   "102_Pilot_Burner_DB_FD_VRFCTN_TMR_ET" : Time = PLC "102_Pilot_Burner_DB".FD_VRFCTN_TMR.ET, 1 s
   "102_Pilot_Burner_DB_FD_VRFCTN_TMR II_ET" : Time = PLC "20_TANKS_IP_DATA".RIO_02.SECOND_TANK.BWT_DO, 1 s
   "86_Times_PIT358 Delay" : Time = PLC "86_Times"."PIT358 Delay", 1 s
   "86_Times_PIT348 Delay" : Time = PLC "86_Times"."PIT348 Delay", 1 s
   "PGC Flush_DB_Temperature Setpoint" : Real = PLC "PGC Flush_DB"."Temperature Setpoint", 1 s
   "2062_Warning_Data_Water Level Override" : Bool = PLC "2062_Warning_Data"."Water Level Override" AT %DB2062.DBX376.0, 1 s
   "2062_Warning_Data_Water Level Override_Aux" : Bool = PLC "2062_Warning_Data"."Water Level Override_Aux" AT %DB2062.DBX376.2, 1 s
   "Sequence Times_DB_Boost" : Bool = PLC "Sequence Times_DB".Boost, 1 s
   "86_Times_FS320 delay" : Time = PLC "86_Times"."FS320 delay", 1 s
   "86_Times_FS317 delay" : Time = PLC "86_Times"."FS317 delay", 1 s
   "86_Times_PS101 Alarm Delay" : Time = PLC "86_Times"."PS101 Alarm Delay", 1 s
   "82_To_HMI_FS350 Animation" : Int = PLC "82_To_HMI"."FS350 Animation", 1 s
   "82_To_HMI_FS332 Animation" : Int = PLC "82_To_HMI"."FS332 Animation", 1 s
   "82_To_HMI_P304 Animation" : Int = PLC "82_To_HMI"."P304 Animation", 1 s
   "Sequence Times_DB_Post-Dwell Timer_Q" : Bool = PLC "Sequence Times_DB"."Post-Dwell Timer".Q, 1 s
      on ChangeValue: "TreatmentCycleCompleted"()
   "51_SLAVE_STATUS_MAIN_BURNER_ACTV" : Bool = PLC "51_SLAVE_STATUS".MAIN_BURNER_ACTV AT %DB51.DBX17.5, 1 s
   "Main Burner Animation_DB_Animation" : Int = PLC "Main Burner Animation_DB".Animation, 1 s
   "20_TANKS_IP_DATA_RIO_01_FIRST_TANK_USD FLOW  N" : Real = PLC "20_TANKS_IP_DATA".RIO_01.FIRST_TANK."USD FLOW  N", 1 s
   "20_TANKS_IP_DATA_RIO_01_FIRST_TANK_MBG_FLOW N" : Real = PLC "20_TANKS_IP_DATA".RIO_01.FIRST_TANK."MBG_FLOW N", 1 s
   "20_TANKS_IP_DATA_RIO_01_SECOND_TANK_MBG_FLOW N" : Real = PLC "20_TANKS_IP_DATA".RIO_01.SECOND_TANK."MBG_FLOW N", 1 s
   "20_TANKS_IP_DATA_RIO_01_SECOND_TANK_USD FLOW  N" : Real = PLC "20_TANKS_IP_DATA".RIO_01.SECOND_TANK."USD FLOW  N", 1 s
   "20_TANKS_IP_DATA_RIO_01_THIRD_TANK_MBG_FLOW N" : Real = PLC "20_TANKS_IP_DATA".RIO_01.THIRD_TANK."MBG_FLOW N", 1 s
   "20_TANKS_IP_DATA_RIO_01_THIRD_TANK_USD FLOW  N" : Real = PLC "20_TANKS_IP_DATA".RIO_01.THIRD_TANK."USD FLOW  N", 1 s
   "20_TANKS_IP_DATA_RIO_03_FIRST_TANK_MBG_FLOW N" : Real = PLC "20_TANKS_IP_DATA".RIO_03.FIRST_TANK."MBG_FLOW N", 1 s
   "20_TANKS_IP_DATA_RIO_03_FIRST_TANK_USD FLOW  N" : Real = PLC "20_TANKS_IP_DATA".RIO_03.FIRST_TANK."USD FLOW  N", 1 s
   "20_TANKS_IP_DATA_RIO_03_SECOND_TANK_USD FLOW  N" : Real = PLC "20_TANKS_IP_DATA".RIO_03.SECOND_TANK."USD FLOW  N", 1 s
   "20_TANKS_IP_DATA_RIO_03_SECOND_TANK_MBG_FLOW N" : Real = PLC "20_TANKS_IP_DATA".RIO_03.SECOND_TANK."MBG_FLOW N", 1 s
   "20_TANKS_IP_DATA_RIO_04_FIRST_TANK_MBG_FLOW N" : Real = PLC "20_TANKS_IP_DATA".RIO_04.FIRST_TANK."MBG_FLOW N", 1 s
   "20_TANKS_IP_DATA_RIO_04_FIRST_TANK_USD FLOW  N" : Real = PLC "20_TANKS_IP_DATA".RIO_04.FIRST_TANK."USD FLOW  N", 1 s
   "20_TANKS_IP_DATA_RIO_04_SECOND_TANK_USD FLOW  N" : Real = PLC "20_TANKS_IP_DATA".RIO_04.SECOND_TANK."USD FLOW  N", 1 s
   "20_TANKS_IP_DATA_RIO_04_SECOND_TANK_MBG_FLOW N" : Real = PLC "20_TANKS_IP_DATA".RIO_04.SECOND_TANK."MBG_FLOW N", 1 s
   "20_TANKS_IP_DATA_RIO_05_FIRST_TANK_MBG_FLOW N" : Real = PLC "20_TANKS_IP_DATA".RIO_05.FIRST_TANK."MBG_FLOW N", 1 s
   "20_TANKS_IP_DATA_RIO_05_FIRST_TANK_USD FLOW  N" : Real = PLC "20_TANKS_IP_DATA".RIO_05.FIRST_TANK."USD FLOW  N", 1 s
   "20_TANKS_IP_DATA_RIO_05_SECOND_TANK_USD FLOW  N" : Real = PLC "20_TANKS_IP_DATA".RIO_05.SECOND_TANK."USD FLOW  N", 1 s
   "20_TANKS_IP_DATA_RIO_05_SECOND_TANK_MBG_FLOW N" : Real = PLC "20_TANKS_IP_DATA".RIO_05.SECOND_TANK."MBG_FLOW N", 1 s
   "20_TANKS_IP_DATA_RIO_06_FIRST_TANK_MBG_FLOW N" : Real = PLC "20_TANKS_IP_DATA".RIO_06.FIRST_TANK."MBG_FLOW N", 1 s
   "20_TANKS_IP_DATA_RIO_06_FIRST_TANK_USD FLOW  N" : Real = PLC "2062_Warning_Data"."Alarm Tank S2", 1 s
   "20_TANKS_IP_DATA_RIO_06_SECOND_TANK_USD FLOW  N" : Real = PLC "86_Times".P304_STRTD_DLY, 1 s
   "20_TANKS_IP_DATA_RIO_06_SECOND_TANK_MBG_FLOW N" : Real = PLC "20_TANKS_IP_DATA".RIO_06.SECOND_TANK."MBG_FLOW N", 1 s
   "20_TANKS_IP_DATA_RIO_07_FIRST_TANK_MBG_FLOW N" : Real = PLC "20_TANKS_IP_DATA".RIO_07.FIRST_TANK."MBG_FLOW N", 1 s
   "20_TANKS_IP_DATA_RIO_07_FIRST_TANK_USD FLOW  N" : Real = PLC "20_TANKS_IP_DATA".RIO_07.FIRST_TANK."USD FLOW  N", 1 s
   "Nm³/hr to m³/hr" : Bool = PLC "80_From_HMI"."m³/hr to Nm³/hr" AT %DB1.DBX0.0, 1 s
   "Ful Pump Ani Animation_DB_Animation" : Int = PLC "Ful Pump Ani Animation_DB".Animation, 1 s
   "IDB_E500B_Animation_Animation" : Int = PLC IDB_E500B_Animation.Animation, 1 s
   "IDB_E500A_Animation_Animation" : Int = PLC IDB_E500A_Animation.Animation, 1 s
   "IDB_E131_Animation_Animation" : Int = PLC IDB_E131_Animation.Animation, 1 s
   "2062_Warning_Data_BTCS_WARNING_WORD_17" : Word = PLC "2062_Warning_Data".BTCS_WARNING_WORD_17 AT %DB2062.DBW372, 1 s
   "IGG HMI HEART BEAT" : Bool = PLC "59_COMMS_HEALTH_DATA"."IGG HMI HB" AT %DB1.DBX0.0, 1 s
   "TRUE" : Bool = PLC AlwaysTRUE AT %M1.2, 1 s
   "IGG PLC HEART BEAT" : Bool = PLC "55_STATUS_DATA".HEART_BEAT AT %DB55.DBX0.0, 100 ms
      on ChangeValue: "HeartBeatFunction"()
   "LOG IGG_1" : Bool = PLC "68_Sys_Status_Data"."LOG IGG" AT %DB1.DBX0.0, 1 s
      on ChangeValue: function_fd9437ed(0, "IGG_IG_TX-431_Atm Oxygen 2"); function_fd9437ed(0, "IGG_CAB_E139_Amps"); function_fd9437ed(0, "CA Blower Pressure Scaled"); function_fd9437ed(0, "IGG_CAB_E139_Comb Air Blower (RPM)"); function_fd9437ed(0, "IGG_IG_CV403_Vent Valve Position"); function_fd9437ed(0, "IGG_BC_FD001_Flame Detector"); function_fd9437ed(0, "IGG_CAB_E139_Setpoint (RPM)"); function_fd9437ed(0, "IGG_IG_TX-600_O2 Setpoint"); function_fd9437ed(0, "IGG_IG_TX-700_Soot Monitor"); function_fd9437ed(0, "IGG_IA_CV111_Atom Air to MBurner-Valve Position"); function_fd9437ed(0, "IGG_IG_TX-600_Oxygen Analyser")
   "LOG GCU" : Bool = PLC "68_Sys_Status_Data"."LOG GCU", 1 s
      on ChangeValue: function_fd9437ed(0, "GCU_IG_TIT406_Gas to deck"); function_fd9437ed(0, "GCU_FW_TIT408_Fresh water cooling"); function_fd9437ed(0, "GCU_SW_PIT348_Sea water cooling"); function_fd9437ed(0, "GCU_FW_PIT353_Fresh water cooling"); function_fd9437ed(0, "GCU_FW_PIT358_Fresh water fill"); function_fd9437ed(0, "GCU_IG_PIT416_Gas to deck"); function_fd9437ed(0, "GCU_Setpoints_PIT416_Target"); function_fd9437ed(0, "PGC_PG_PT002_PGC Outlet"); function_fd9437ed(0, "PGC_PG_TE002_PGC Outlet"); function_fd9437ed(0, "GCU_FW_LIT304_GCU Level"); function_fd9437ed(0, "GCU_SL_400_SCALED"); function_fd9437ed(0, "BWT_Setpoints_DO_SP"); function_fd9437ed(0, "GCU_FW_LIT305_IBC Tank Level"); function_fd9437ed(0, "BWT_2P_FIT-420_MBG Flow_Raw"); function_fd9437ed(0, "BWT_2P_FIT-418_USD Flow_Raw"); function_fd9437ed(0, "BWT_2S_FIT-419_MBG Flow_Raw")
   "LOG GCU_1" : Bool = PLC "68_Sys_Status_Data"."LOG GCU", 1 s
      on ChangeValue: function_fd9437ed(0, "BWT_2S_FIT-417_USD Flow_Raw"); function_fd9437ed(0, "Treatment check"); function_fd9437ed(0, "BWT_3P"); function_fd9437ed(0, "BWT_3S"); function_fd9437ed(0, "BWT_4P"); function_fd9437ed(0, "BWT_4S"); function_fd9437ed(0, "BWT_5P"); function_fd9437ed(0, "BWT_5S"); function_fd9437ed(0, "BWT_6P"); function_fd9437ed(0, "BWT_6S"); function_fd9437ed(0, "BWT APT"); function_fd9437ed(0, "BWT_2P"); function_fd9437ed(0, "BWT_2S"); function_fd9437ed(0, "BWT_1P"); function_fd9437ed(0, "BWT_FPT"); function_fd9437ed(0, "BWT_1S")
   "LOG GCU_2" : Bool = PLC "68_Sys_Status_Data"."LOG GCU", 1 s
      on ChangeValue: function_fd9437ed(0, "GCU_CV405_Vent Valve Position")
   "STOP LOG GCU" : Bool = PLC "68_Sys_Status_Data"."STOP LOG GCU" AT %DB1.DBX0.0, 1 s
      on ChangeValue: function_b6526003(0, "GCU_IG_TIT406_Gas to deck"); function_b6526003(0, "GCU_FW_TIT408_Fresh water cooling"); function_b6526003(0, "GCU_SW_PIT348_Sea water cooling"); function_b6526003(0, "GCU_FW_PIT353_Fresh water cooling"); function_b6526003(0, "GCU_FW_PIT358_Fresh water fill"); function_b6526003(0, "GCU_IG_PIT416_Gas to deck"); function_b6526003(0, "GCU_Setpoints_PIT416_Target"); function_b6526003(0, "PGC_PG_PT002_PGC Outlet"); function_b6526003(0, "PGC_PG_TE002_PGC Outlet"); function_b6526003(0, "GCU_FW_LIT304_GCU Level"); function_b6526003(0, "GCU_SL_400_SCALED"); function_b6526003(0, "BWT_Setpoints_DO_SP"); function_b6526003(0, "GCU_FW_LIT305_IBC Tank Level"); function_b6526003(0, "BWT_2P_FIT-420_MBG Flow_Raw"); function_b6526003(0, "BWT_2P_FIT-418_USD Flow_Raw"); function_b6526003(0, "BWT_2S_FIT-419_MBG Flow_Raw")
   "STOP LOG IGG" : Bool = PLC "68_Sys_Status_Data"."STOP LOG IGG" AT %DB1.DBX0.0, 1 s
      on ChangeValue: function_b6526003(0, "IGG_Fuel_TIT202_Fuel Oil"); function_b6526003(0, "IGG_IG_TIT401_IG vent"); function_b6526003(0, "IGG_SW_TIT319_Cooling water (main line)"); function_b6526003(0, "IGG_SW_TIT360_Cooling water to drain line"); function_b6526003(0, "IGG_SW_TIT315_CW Temp to IGG Jacket"); function_b6526003(0, "IGG_CAB_PIT102_Comb Air"); function_b6526003(0, "IGG_Fuel_PIT204_Fuel Oil"); function_b6526003(0, "IGG_IA_PIT113_Atom Air to MBurner"); function_b6526003(0, "IGG_Fuel_PIT205_Fuel to MBurner"); function_b6526003(0, "IGG_IG_PIT402_IG vent"); function_b6526003(0, "IGG_SW_PIT359_Cooling water (main line)"); function_b6526003(0, "IGG_IA_PIT112_Inst Air"); function_b6526003(0, "IGG_SW_PIT316_Cooling water to IGG Jacket"); function_b6526003(0, "IGG_IG_TX-431_Atm Oxygen 1"); function_b6526003(0, "IGG_IG_TX-431_Atm Oxygen 2"); function_b6526003(0, "IGG_CAB_E139_Amps")
   "STOP LOG GCU_1" : Bool = PLC "68_Sys_Status_Data"."STOP LOG GCU" AT %DB1.DBX0.0, 1 s
      on ChangeValue: function_b6526003(0, "BWT_2S_FIT-417_USD Flow_Raw"); function_b6526003(0, "BWT_3P"); function_b6526003(0, "BWT_3S"); function_b6526003(0, "BWT_4P"); function_b6526003(0, "BWT_4S"); function_b6526003(0, "BWT_5P"); function_b6526003(0, "BWT_5S"); function_b6526003(0, "BWT_6P"); function_b6526003(0, "BWT_6S"); function_b6526003(0, "BWT APT"); function_b6526003(0, "BWT_2P"); function_b6526003(0, "BWT_2S"); function_b6526003(0, "BWT_1P"); function_b6526003(0, "BWT_FPT"); function_b6526003(0, "BWT_1S"); function_b6526003(0, "GCU_CV405_Vent Valve Position")
   "STOP LOG IGG_1" : Bool = PLC "68_Sys_Status_Data"."STOP LOG IGG" AT %DB1.DBX0.0, 1 s
      on ChangeValue: function_b6526003(0, "IGG_CAB_E139_Comb Air Blower (RPM)"); function_b6526003(0, "IGG_IG_CV403_Vent Valve Position"); function_b6526003(0, "IGG_BC_FD001_Flame Detector"); function_b6526003(0, "IGG_CAB_E139_Setpoint (RPM)"); function_b6526003(0, "IGG_IG_TX-600_O2 Setpoint"); function_b6526003(0, "IGG_IG_TX-700_Soot Monitor"); function_b6526003(0, "IGG_IA_CV111_Atom Air to MBurner-Valve Position"); function_b6526003(0, "IGG_IG_TX-600_Oxygen Analyser")
   "HEART BEAT TRUE" : Bool = PLC "68_Sys_Status_Data"."TRUE for HMI" AT %M1.2, 100 ms
   "80_From_HMI_Jurney Start Simulator" : Bool = PLC "80_From_HMI"."Jurney Start Simulator", 1 s
   "68_Sys_Status_Data_LOG IGG Simulator" : Bool = PLC "68_Sys_Status_Data"."LOG IGG Simulator", 1 s
   "68_Sys_Status_Data_LOG GCU Simulator" : Bool = PLC "68_Sys_Status_Data"."LOG GCU Simulator", 1 s
   "Setpoint Override_DB_Activate Press Prot" : Bool = PLC "Setpoint Override_DB"."Activate Press Prot", 1 s
   "Setpoint Override_DB_Temperature Tolerance" : Real = PLC "Setpoint Override_DB"."Temperature Tolerance", 1 s
   "Setpoint Override_DB_Pressure Tolerance" : Real = PLC "Setpoint Override_DB"."Pressure Tolerance", 1 s
   "Setpoint Override_DB_Activate Temp Prot" : Bool = PLC "Setpoint Override_DB"."Activate Temp Prot", 1 s
   "Setpoint Override_DB_Reset" : Bool = PLC "Setpoint Override_DB".Reset, 1 s
   "Setpoint Override_DB_Tank Change TimeOut" : Time = PLC "Setpoint Override_DB"."Tank Change TimeOut", 1 s
   "Setpoint Override_DB_Set Pressure" : Bool = PLC "Setpoint Override_DB"."Set Pressure", 1 s
      on ChangeValue: function_efd93a16("PGC Protection Warning", 300, 200, -1, 3, 1)
   "80_From_HMI_TT002 Target Protection" : Bool = PLC "80_From_HMI"."TT002 Target Protection", 1 s
   "80_From_HMI_PT002 Target Protection" : Bool = PLC "80_From_HMI"."PT002 Target Protection", 1 s
   "80_From_HMI_Tank Close Protection" : Bool = PLC "80_From_HMI"."Tank Close Protection", 1 s
   "84_Setpoints_PIT416_Target_Safe" : Real = PLC "84_Setpoints".PIT416_Target_Safe, 1 s
   "84_Setpoints_Tank Close TimeOut" : Time = PLC "84_Setpoints"."Tank Close TimeOut", 1 s
   "84_Setpoints_E-400 PT002 Tolerance" : Real = PLC "84_Setpoints"."E-400 PT002 Tolerance", 1 s
   "84_Setpoints_E-400 TT002 Tolerance" : Real = PLC "84_Setpoints"."E-400 TT002 Tolerance", 1 s
   "Sequence Times_DB_Jurney Timer_Days Left" : DInt = PLC "Sequence Times_DB"."Jurney Timer"."Days Left", 1 s
   "Sequence Times_DB_Jurney Timer_Hours Left" : DInt = PLC "Sequence Times_DB"."Jurney Timer"."Hours Left", 1 s
   "Sequence Times_DB_Jurney Timer_Minutes Left" : DInt = PLC "Sequence Times_DB"."Jurney Timer"."Minutes Left", 1 s
   "2086_Times_Stage Warning" : Time = PLC "2062_Warning_Data"."Water Level Override 1S", 1 s
   "Warn To Start IGG" : Bool = PLC "82_To_HMI"."Warn to Start IGG", 1 s
      on ChangeValue: "TimeRemainingToTreatment"()
   "Warn To Start IGG-Last" : Bool = PLC "82_To_HMI"."Warn to Start IGG-Last", 1 s
      on ChangeValue: "TreatmentRequired"()
   "Warn To Start GCU" : Bool = PLC "82_To_HMI"."Warn to Start GCU", 1 s
      on ChangeValue: "TimeRemainingToRe_Ox"()
   "Warn To Start GCU-Last" : Bool = PLC "82_To_HMI"."Warn to Start GCU-Last", 1 s
      on ChangeValue: "TreatmentRequired_GCU"()
   "80_From_HMI_GCU Start Confirmed" : Bool = PLC "80_From_HMI"."GCU Start Confirmed", 1 s
      on ChangeValue: "TreatmentRequired_GCU"()
   "102_Pilot_Burner_DB_STATE" : Int = PLC "102_Pilot_Burner_DB".STATE, 1 s
   "Tag_1" : Bool = PLC Tag_1 AT %M233.3, 1 s
   "Tag_2" : Bool = PLC Tag_2 AT %M233.4, 1 s
   "Tag_3" : Bool = PLC Tag_3 AT %M233.5, 1 s
   "Tag_4" : Bool = PLC Tag_4 AT %M233.6, 1 s
   "Tag_5" : Bool = PLC Tag_5 AT %M233.7, 1 s
   "2068_Sys_Status_Data_Times Visibil" : Bool = PLC "2068_Sys_Status_Data"."Times Visibil", 1 s
   "Sequence Times_DB_Warn to GCU Start" : Bool = PLC "Sequence Times_DB"."Warn to GCU Start", 1 s
   "80_From_HMI_CSW OVR Stop" : Bool = PLC "80_From_HMI"."CSW OVR Stop", 1 s
   "Sequence Times_DB_Offset Timer_Days Left" : DInt = PLC "Sequence Times_DB"."Offset Timer"."Days Left", 1 s
   "Sequence Times_DB_Offset Timer_Hours Left" : DInt = PLC "Sequence Times_DB"."Offset Timer"."Hours Left", 1 s
   "Sequence Times_DB_Offset Timer_Minutes Left" : DInt = PLC "Sequence Times_DB"."Offset Timer"."Minutes Left", 1 s
   "Voyage Time Invalid" : Bool = PLC "Sequence Times_DB"."Voiage Time Invalid" AT %DB1.DBX0.0, 1 s
      on ChangeValue: "VoyageTimeInsufficient"()
   "82_To_HMI_IGG RUN Indication" : Bool = PLC "82_To_HMI"."IGG RUN Indication", 1 s
   "Not TANK Activ Warning" : Bool = PLC "2068_Sys_Status_Data"."Not TANK Activ Warning" AT %DB1.DBX0.0, 1 s
      on ChangeValue: "TANK_Activ_Warning"()
   "Sequence Times_DB_Pre-Dwell Done" : Bool = PLC "Sequence Times_DB"."Pre-Dwell Done", 1 s
   "Sequence Times_DB_De-Ox Done" : Bool = PLC "Sequence Times_DB"."De-Ox Done", 1 s
   "Sequence Times_DB_Dwell Done" : Bool = PLC "Sequence Times_DB"."Dwell Done", 1 s
   "Sequence Times_DB_Re-Ox Done" : Bool = PLC "Sequence Times_DB"."Re-Ox Done", 1 s
   "Sequence Times_DB_Post-Dwell Done" : Bool = PLC "Sequence Times_DB"."Post-Dwell Done", 1 s

HMI tags "Alarms"
   "60_Alarm_Data_BC_ALARM_WORD_01" : Word = PLC "60_Alarm_Data".BC_ALARM_WORD_01 AT %DB60.DBW0, 1 s
   "60_Alarm_Data_BC_ALARM_WORD_02" : Word = PLC "60_Alarm_Data".BC_ALARM_WORD_02 AT %DB60.DBW2, 1 s
   "60_Alarm_Data_BC_ALARM_WORD_03" : Word = PLC "60_Alarm_Data".BC_ALARM_WORD_03 AT %DB60.DBW4, 1 s
   "60_Alarm_Data_BC_ALARM_WORD_04" : Word = PLC "60_Alarm_Data".BC_ALARM_WORD_04 AT %DB60.DBW6, 1 s
   "60_Alarm_Data_GCU_ALARM_WORD_01" : Word = PLC "60_Alarm_Data".GCU_ALARM_WORD_01 AT %DB60.DBW0, 1 s
   "60_Alarm_Data_GCU_ALARM_WORD_02" : Word = PLC "60_Alarm_Data".GCU_ALARM_WORD_02 AT %DB60.DBW2, 1 s
   "60_Alarm_Data_GCU_ALARM_WORD_03" : Word = PLC "60_Alarm_Data".GCU_ALARM_WORD_03 AT %DB60.DBW4, 1 s
   "60_Alarm_Data_GCU_ALARM_WORD_04" : Word = PLC "60_Alarm_Data".GCU_ALARM_WORD_04 AT %DB60.DBW6, 1 s
   "60_Alarm_Data_GCU_ALARM_WORD_05" : Word = PLC "60_Alarm_Data".GCU_ALARM_WORD_05 AT %DB60.DBW8, 1 s
   "60_Alarm_Data_GCU_ALARM_WORD_06" : Word = PLC "60_Alarm_Data".GCU_ALARM_WORD_06 AT %DB60.DBW10, 1 s
   "60_Alarm_Data_GCU_ALARM_WORD_07" : Word = PLC "60_Alarm_Data".GCU_ALARM_WORD_07 AT %DB60.DBW12, 1 s
   "60_Alarm_Data_GCU_ALARM_WORD_08" : Word = PLC "60_Alarm_Data".GCU_ALARM_WORD_08 AT %DB60.DBW14, 1 s
   "60_Alarm_Data_GCU_ALARM_WORD_09" : Word = PLC "60_Alarm_Data".GCU_ALARM_WORD_09 AT %DB60.DBW16, 1 s
   "60_Alarm_Data_IGG_ALARM_WORD_01" : Word = PLC "60_Alarm_Data".IGG_ALARM_WORD_01 AT %DB60.DBW0, 1 s
   "60_Alarm_Data_IGG_ALARM_WORD_02" : Word = PLC "60_Alarm_Data".IGG_ALARM_WORD_02 AT %DB60.DBW2, 1 s
   "60_Alarm_Data_IGG_ALARM_WORD_03" : Word = PLC "60_Alarm_Data".IGG_ALARM_WORD_03 AT %DB60.DBW4, 1 s
   "60_Alarm_Data_IGG_ALARM_WORD_04" : Word = PLC "60_Alarm_Data".IGG_ALARM_WORD_04 AT %DB60.DBW6, 1 s
   "2060_Alarm_Data_BTCS_ALARM_WORD_01" : Word = PLC "2060_Alarm_Data".BTCS_ALARM_WORD_01 AT %DB2060.DBW0, 1 s
   "2060_Alarm_Data_BTCS_ALARM_WORD_02" : Word = PLC "2060_Alarm_Data".BTCS_ALARM_WORD_02 AT %DB2060.DBW2, 1 s
   "2060_Alarm_Data_BTCS_ALARM_WORD_03" : Word = PLC "2060_Alarm_Data".BTCS_ALARM_WORD_03 AT %DB2060.DBW4, 1 s
   "2060_Alarm_Data_BTCS_ALARM_WORD_04" : Word = PLC "2060_Alarm_Data".BTCS_ALARM_WORD_04 AT %DB2060.DBW6, 1 s
   "2060_Alarm_Data_BTCS_ALARM_WORD_05" : Word = PLC "2060_Alarm_Data".BTCS_ALARM_WORD_05 AT %DB2060.DBW8, 1 s
   "2060_Alarm_Data_BTCS_ALARM_WORD_06" : Word = PLC "2060_Alarm_Data".BTCS_ALARM_WORD_06 AT %DB2060.DBW10, 1 s
   "2060_Alarm_Data_BTCS_ALARM_WORD_07" : Word = PLC "2060_Alarm_Data".BTCS_ALARM_WORD_07 AT %DB2060.DBW12, 1 s
   "2060_Alarm_Data_BTCS_ALARM_WORD_08" : Word = PLC "2060_Alarm_Data".BTCS_ALARM_WORD_08 AT %DB2060.DBW14, 1 s

HMI tags "BC_HMI_Tags"
   "10 DI_DATA_E131_OK" : Bool = PLC "20_TANKS_IP_DATA".RIO_03.FIRST_TANK.USD_FLOW AT %DB1.DBX0.0, 1 s
   "10 DI_DATA_E131_SHTDN" : Bool = PLC "10 DI_DATA".E131_SHTDN AT %DB1.DBX0.0, 1 s
   "103_Main_Burner_DB_DN_OK(1)" : Bool = PLC "103_Main_Burner_DB".DN_OK AT %DB1.DBX0.0, 1 s
   "10 DI_DATA_FD001_OK" : Bool = PLC "10 DI_DATA".FD001_OK AT %DB1.DBX0.0, 1 s
   "10 DI_DATA_FD001_PWR_OK" : Bool = PLC "10 DI_DATA".FD001_PWR_OK AT %DB1.DBX0.0, 1 s
   "10 DI_DATA_FS115(1)" : Bool = PLC "10 DI_DATA".FS115 AT %DB1.DBW0, 1 s
   "10 DI_DATA_FS123" : Bool = PLC "10 DI_DATA".FS123 AT %DB1.DBX0.0, 1 s
   "10 DI_DATA_FS317" : Bool = PLC "10 DI_DATA".FS317 AT %DB1.DBX0.0, 1 s
   "10 DI_DATA_FS320" : Bool = PLC "10 DI_DATA".FS320 AT %DB1.DBX0.0, 1 s
   "10 DI_DATA_ESD_OK" : Bool = PLC "10 DI_DATA".ESD_OK AT %DB1.DBX0.0, 1 s
   "10 DI_DATA_P301_ENBLD" : Bool = PLC "10 DI_DATA".P301_ENBLD AT %DB1.DBX0.0, 1 s
   "10 DI_DATA_R2_SPR_DI_1_6" : Bool = PLC "10 DI_DATA".R2_SPR_DI_1_6 AT %DB1.DBX0.0, 1 s
   "10 DI_DATA_P301_TRIPPED(1)" : Bool = PLC "10 DI_DATA".P301_TRIPPED AT %DB1.DBX0.0, 1 s
   "10 DI_DATA_P305_ENBLD" : Bool = PLC "10 DI_DATA".P305_ENBLD AT %DB1.DBX0.0, 1 s
   "10 DI_DATA_P305_TRIPPED(1)" : Bool = PLC "10 DI_DATA".P305_TRIPPED AT %DB1.DBX0.0, 1 s
   "10 DI_DATA_PS101" : Bool = PLC "10 DI_DATA".PS101 AT %DB1.DBX0.0, 1 s
   "10 DI_DATA_R2_SPR_DI_0_2" : Bool = PLC "10 DI_DATA".R2_SPR_DI_0_2 AT %DB1.DBX0.0, 1 s
   "10 DI_DATA_R2_SPR_DI_0_3" : Bool = PLC "10 DI_DATA".R2_SPR_DI_0_3 AT %DB1.DBX0.0, 1 s
   "10 DI_DATA_TS403_FAULT" : Bool = PLC "10 DI_DATA".TS403_FAULT AT %DB1.DBX0.0, 1 s
   "10 DI_DATA_X001_PWR_OK" : Bool = PLC "10 DI_DATA".X001_PWR_OK AT %DB1.DBX0.0, 1 s
   "102_Pilot_Burner_DB_FLM_DET" : Bool = PLC "102_Pilot_Burner_DB".FLM_DET AT %DB1.DBX0.0, 100 ms
   "104_Pilot_Purge_DB_DN_OK" : Bool = PLC "104_Pilot_Purge_DB".DN_OK AT %DB1.DBX0.0, 1 s
   "10 DI_DATA_E600_NOK" : Bool = PLC "10 DI_DATA".E600_NOK AT %DB1.DBX0.0, 1 s
   "10 DI_DATA_E600_HIHI" : Bool = PLC "10 DI_DATA".E600_HIHI AT %DB1.DBX0.0, 1 s
   "10 DI_DATA_E600_LOLO" : Bool = PLC "10 DI_DATA".E600_LOLO AT %DB1.DBX0.0, 1 s
   "10 DI_DATA_E600_PWR_OK" : Bool = PLC "10 DI_DATA".E600_PWR_OK AT %DB1.DBX0.0, 1 s
   "10 DI_DATA_E700_PWR_OK" : Bool = PLC "10 DI_DATA".E700_PWR_OK AT %DB1.DBX0.0, 1 s
   "10 DI_DATA_E700_OPACITY" : Bool = PLC "10 DI_DATA".E700_OPACITY AT %DB1.DBX0.0, 1 s
   "10 DI_DATA_TS403_FAULT(1)" : Bool = PLC "10 DI_DATA".TS403_FAULT AT %DB1.DBX0.0, 1 s
   "10 DI_DATA_TS006" : Bool = PLC "10 DI_DATA".TS006 AT %DB1.DBX0.0, 1 s
   "10 DI_DATA_S2_8K1_OK" : Bool = PLC "10 DI_DATA".S2_8K1_OK AT %DB1.DBX0.0, 1 s
   "10 DI_DATA_E131_WRNG" : Bool = PLC "10 DI_DATA".E131_WRNG AT %DB1.DBX0.0, 1 s
   "10 DI_DATA_R2_SPR_DI_3_2" : Bool = PLC "10 DI_DATA".R2_SPR_DI_3_2 AT %DB1.DBX0.0, 1 s
   "10 DI_DATA_R2_SPR_DI_3_7" : Bool = PLC "10 DI_DATA".R2_SPR_DI_3_7 AT %DB1.DBX0.0, 1 s
   "10 DI_DATA_LS001" : Bool = PLC "10 DI_DATA".LS001 AT %DB1.DBX0.0, 1 s
   "10 DI_DATA_P305_TRIPPED" : Bool = PLC "10 DI_DATA".P305_TRIPPED AT %DB1.DBX0.0, 1 s
   "10 DI_DATA_P305_ENBLD(1)" : Bool = PLC "10 DI_DATA".P305_ENBLD AT %DB1.DBX0.0, 1 s
   "84_Setpoints_PIT113_High" : Real = PLC "84_Setpoints".PIT113_High AT %DB1.DBD0, 1 s
   "84_Setpoints_PIT113_HighHigh" : Real = PLC "84_Setpoints".PIT113_HighHigh AT %DB1.DBD0, 1 s
   "84_Setpoints_PIT113_Pilot_Target" : Real = PLC "84_Setpoints".PIT113_Pilot_Target AT %DB1.DBX0.0, 1 s
   "84_Setpoints_PIT204_High(2)" : Real = PLC "84_Setpoints".PIT204_High, 1 s
   "84_Setpoints_PIT204_HighHigh(2)" : Real = PLC "84_Setpoints".PIT204_HighHigh, 1 s
   "84_Setpoints_PIT204_Low(2)" : Real = PLC "84_Setpoints".PIT204_Low, 1 s
   "84_Setpoints_PIT204_LowLow(2)" : Real = PLC "84_Setpoints".PIT204_LowLow, 1 s
   "84_Setpoints_PIT205_High" : Real = PLC "2084_Setpoints"."TX427 Star DO Lo" AT %DB1.DBD0, 1 s
   "84_Setpoints_PIT205_HighHigh" : Real = PLC "84_Setpoints".PIT205_HighHigh AT %DB1.DBD0, 1 s
   "84_Setpoints_PIT205_Low" : Real = PLC "84_Setpoints".PIT205_Low AT %DB1.DBD0, 1 s
   "84_Setpoints_PIT205_LowLow" : Real = PLC "84_Setpoints".PIT205_LowLow AT %DB1.DBD0, 1 s
   "84_Setpoints_PIT205_Target" : Real = PLC "84_Setpoints".PIT205_Target AT %DB1.DBX0.0, 1 s
   "84_Setpoints_PIT113_Low" : Real = PLC "84_Setpoints".PIT113_Low AT %DB1.DBD0, 1 s
   "84_Setpoints_PIT113_LowLow" : Real = PLC "84_Setpoints".PIT113_LowLow AT %DB1.DBD0, 1 s
   "84_Setpoints_TIT202_High" : Real = PLC "84_Setpoints".TIT202_High AT %DB1.DBD0, 1 s
   "84_Setpoints_TIT202_HighHigh" : Real = PLC "84_Setpoints".TIT202_HighHigh AT %DB1.DBD0, 1 s
   "84_Setpoints_TIT202_LowLow" : Real = PLC "84_Setpoints".TIT202_LowLow AT %DB1.DBD0, 1 s
   "84_Setpoints_TIT202_Low" : Real = PLC "84_Setpoints".TIT202_Low AT %DB1.DBD0, 1 s
   "84_Setpoints_TX700_High" : Real = PLC "84_Setpoints".TX700_High AT %DB1.DBD0, 1 s
   "84_Setpoints_TX700_Low" : Real = PLC "84_Setpoints".TX700_Low AT %DB1.DBD0, 1 s
   "84_Setpoints_FD001_LowLow" : Real = PLC "84_Setpoints".FD001_LowLow AT %DB1.DBD0, 1 s
   "84_Setpoints_E600_BWT_High" : Real = PLC "84_Setpoints".E600_BWT_High AT %DB1.DBD0, 1 s
   "84_Setpoints_E600_BWT_Low" : Real = PLC "84_Setpoints".E600_BWT_Low AT %DB1.DBD0, 1 s
   "84_Setpoints_FD001_Low" : Real = PLC "84_Setpoints".FD001_Low AT %DB1.DBD0, 1 s
   "84_Setpoints_AT_O2_1_LowLow" : Real = PLC "84_Setpoints".AT_O2_1_LowLow AT %DB1.DBD0, 1 s
   "84_Setpoints_AT_O2_2_LowLow" : Real = PLC "84_Setpoints".AT_O2_2_LowLow AT %DB1.DBD0, 1 s
   "84_Setpoints_AT_O2_2_Low" : Real = PLC "84_Setpoints".AT_O2_2_Low AT %DB1.DBD0, 1 s
   "80_From_HMI_MAN_DQ_1_7(1)" : Bool = PLC "80_From_HMI".MAN_DQ_1_7 AT %DB1.DBX0.0, 1 s
   "80_From_HMI_MAN_DQ_1_6" : Bool = PLC "80_From_HMI".MAN_DQ_1_6 AT %DB1.DBX0.0, 1 s
   "80_From_HMI_MAN_DQ_1_5(1)" : Bool = PLC "80_From_HMI".MAN_DQ_1_5 AT %DB1.DBX0.0, 1 s
   "80_From_HMI_MAN_DQ_1_4(1)" : Bool = PLC "80_From_HMI".MAN_DQ_1_4 AT %DB1.DBX0.0, 1 s
   "80_From_HMI_MAN_DQ_1_3(1)" : Bool = PLC "80_From_HMI".MAN_DQ_1_3 AT %DB1.DBX0.0, 1 s
   "80_From_HMI_MAN_DQ_1_2(1)" : Bool = PLC "80_From_HMI".MAN_DQ_1_2 AT %DB1.DBX0.0, 1 s
   "80_From_HMI_MAN_DQ_1_1(1)" : Bool = PLC "80_From_HMI".MAN_DQ_1_1 AT %DB1.DBX0.0, 1 s
   "80_From_HMI_MAN_DQ_1_0" : Bool = PLC "80_From_HMI".MAN_DQ_1_0 AT %DB1.DBX0.0, 1 s
   "80_From_HMI_MAN_DQ_0_7" : Bool = PLC "80_From_HMI".MAN_DQ_0_7 AT %DB1.DBX0.0, 1 s
   "80_From_HMI_MAN_DQ_0_6(1)" : Bool = PLC "80_From_HMI".MAN_DQ_0_6 AT %DB1.DBX0.0, 1 s
   "80_From_HMI_MAN_DQ_0_5(1)" : Bool = PLC "80_From_HMI".MAN_DQ_0_5 AT %DB1.DBX0.0, 1 s
   "80_From_HMI_MAN_DQ_0_4(1)" : Bool = PLC "80_From_HMI".MAN_DQ_0_4 AT %DB1.DBX0.0, 1 s
   "80_From_HMI_MAN_DQ_0_3(1)" : Bool = PLC "80_From_HMI".MAN_DQ_0_3 AT %DB1.DBX0.0, 1 s
   "80_From_HMI_MAN_DQ_0_2(1)" : Bool = PLC "80_From_HMI".MAN_DQ_0_2 AT %DB1.DBX0.0, 1 s
   "80_From_HMI_MAN_DQ_0_1(1)" : Bool = PLC "80_From_HMI".MAN_DQ_0_1 AT %DB1.DBX0.0, 1 s
   "80_From_HMI_MAN_DQ_0_0(1)" : Bool = PLC "80_From_HMI".MAN_DQ_0_0 AT %DB1.DBX0.0, 1 s
   "16_AQ_Data_CV111_CNTRL" : Real = PLC "16_AQ_Data".CV111_CNTRL AT %DB1.DBD0, 1 s
   "14_DQ_Data_X001ControlOut" : Bool = PLC "14_DQ_Data".X001ControlOut AT %DB1.DBX0.0, 1 s
   "14_DQ_Data_R2_SPR_DQ_1_6" : Bool = PLC "14_DQ_Data".R2_SPR_DQ_1_6 AT %DB1.DBX0.0, 1 s
   "14_DQ_Data_R2_SPR_DQ_1_4" : Bool = PLC "14_DQ_Data".R2_SPR_DQ_1_4 AT %DB1.DBX0.0, 1 s
   "14_DQ_Data_R2_SPR_DQ_1_5" : Bool = PLC "14_DQ_Data".R2_SPR_DQ_1_5 AT %DB1.DBX0.0, 1 s
   "14_DQ_Data_R2_SPR_DQ_1_3" : Bool = PLC "14_DQ_Data".R2_SPR_DQ_1_3 AT %DB1.DBX0.0, 1 s
   "14_DQ_Data_R2_SPR_DQ_1_2" : Bool = PLC "14_DQ_Data".R2_SPR_DQ_1_2 AT %DB1.DBX0.0, 1 s
   "14_DQ_Data_P305ControlOut" : Bool = PLC "14_DQ_Data".P305ControlOut AT %DB1.DBX0.0, 1 s
   "14_DQ_Data_E131ControlOut" : Bool = PLC "14_DQ_Data".E131ControlOut AT %DB1.DBX0.0, 1 s
   "14_DQ_Data_200CV216ControlOut" : Bool = PLC "14_DQ_Data".200CV216ControlOut AT %DB1.DBX0.0, 1 s
   "14_DQ_Data_200CV215ControlOut" : Bool = PLC "14_DQ_Data".200CV215ControlOut AT %DB1.DBX0.0, 1 s
   "14_DQ_Data_200CV207ControlOut" : Bool = PLC "14_DQ_Data".200CV207ControlOut AT %DB1.DBX0.0, 1 s
   "14_DQ_Data_200CV206ControlOut" : Bool = PLC "14_DQ_Data".200CV206ControlOut AT %DB1.DBX0.0, 1 s
   "14_DQ_Data_200CV127ControlOut" : Bool = PLC "14_DQ_Data".200CV127ControlOut AT %DB1.DBX0.0, 1 s
   "14_DQ_Data_200CV124ControlOut" : Bool = PLC "14_DQ_Data".200CV124ControlOut AT %DB1.DBX0.0, 1 s
   "14_DQ_Data_200CV114ControlOut" : Bool = PLC "14_DQ_Data".200CV114ControlOut AT %DB1.DBX0.0, 1 s
   "12_AI_Data_TIT202In_SCALED" : Real = PLC "12_AI_Data".TIT202In_SCALED AT %DB1.DBX0.0, 1 s
   "12_AI_Data_PIT205In_SCALED" : Real = PLC "12_AI_Data".PIT205In_SCALED AT %DB1.DBX0.0, 1 s
   "12_AI_Data_PIT204In_SCALED" : Real = PLC "12_AI_Data".PIT204In_SCALED AT %DB1.DBX0.0, 1 s
   "12_AI_Data_PIT113In_SCALED" : Real = PLC "12_AI_Data".PIT113In_SCALED AT %DB1.DBD0, 1 s
   "12_AI_Data_PIT112In_SCALED" : Real = PLC "12_AI_Data".PIT112In_SCALED AT %DB1.DBX0.0, 1 s
   "12_AI_Data_FD001FlameSignalIn" : Real = PLC "12_AI_Data".FD001FlameSignalIn AT %DB1.DBX0.0, 100 ms
   "12_AI_Data_E700SootContentIn" : Real = PLC "12_AI_Data".E700SootContentIn AT %DB1.DBX0.0, 1 s
   "12_AI_Data_E600O2ContentIn" : Real = PLC "12_AI_Data".E600O2ContentIn AT %DB1.DBX0.0, 100 ms
   "10 DI_DATA_TS403_FAULT(2)" : Bool = PLC "10 DI_DATA".TS403_FAULT AT %DB1.DBX0.0, 1 s
   "10_DI_Data_E139_RUNNING" : Bool = PLC "10_DI_Data".E139_RUNNING AT %DB1.DBX0.0, 1 s
   "10 DI_DATA_TS006(1)" : Bool = PLC "10 DI_DATA".TS006 AT %DB1.DBX0.0, 1 s
   "16_AQ_Data_CV203_CNTRL" : Real = PLC "16_AQ_Data".CV203_CNTRL AT %DB1.DBD0, 1 s
   "16_AQ_Data_R2_SPR_AQ_96" : Real = PLC "16_AQ_Data".R2_SPR_AQ_96 AT %DB1.DBD0, 1 s
   "16_AQ_Data_R2_SPR_AQ_98" : Real = PLC "16_AQ_Data".R2_SPR_AQ_98 AT %DB1.DBD0, 1 s
   "80_From_HMI_MAN_AQ_INC_96" : Bool = PLC "80_From_HMI".MAN_AQ_INC_96 AT %DB1.DBX0.0, 1 s
   "80_From_HMI_MAN_AQ_DEC_96" : Bool = PLC "80_From_HMI".MAN_AQ_DEC_96 AT %DB1.DBX0.0, 1 s
   "80_From_HMI_MAN_AQ_INC_98" : Bool = PLC "80_From_HMI".MAN_AQ_INC_98 AT %DB1.DBX0.0, 1 s
   "80_From_HMI_MAN_AQ_DEC_98" : Bool = PLC "80_From_HMI".MAN_AQ_DEC_98 AT %DB1.DBX0.0, 1 s
   "80_From_HMI_MAN_AQ_INC_100(1)" : Bool = PLC "80_From_HMI".MAN_AQ_INC_100 AT %DB1.DBX0.0, 1 s
   "80_From_HMI_MAN_AQ_DEC_100(1)" : Bool = PLC "80_From_HMI".MAN_AQ_DEC_100 AT %DB1.DBX0.0, 1 s
   "80_From_HMI_MAN_AQ_INC_102" : Bool = PLC "80_From_HMI".MAN_AQ_INC_102 AT %DB1.DBX0.0, 1 s
   "80_From_HMI_MAN_AQ_DEC_102" : Bool = PLC "80_From_HMI".MAN_AQ_DEC_102 AT %DB1.DBX0.0, 1 s
   "10 DI_DATA_FS115" : Bool = PLC "10 DI_DATA".FS115 AT %DB1.DBX0.0, 1 s
   "10 DI_DATA_P301_TRIPPED" : Bool = PLC "10 DI_DATA".P301_TRIPPED AT %DB1.DBX0.0, 1 s
   "84_Setpoints_E600_BWT_HighHigh" : Real = PLC "84_Setpoints".E600_BWT_HighHigh AT %DB1.DBD0, 1 s
   "84_Setpoints_E600_BWT_LowLow" : Real = PLC "84_Setpoints".E600_BWT_LowLow AT %DB1.DBD0, 1 s
   "84_Setpoints_E600_CB_Low" : Real = PLC "84_Setpoints".E600_CB_Low AT %DB1.DBD0, 1 s
   "84_Setpoints_E600_CB_LowLow" : Real = PLC "84_Setpoints".E600_CB_LowLow AT %DB1.DBD0, 1 s
   "84_Setpoints_E600_CB_High" : Real = PLC "84_Setpoints".E600_CB_High AT %DB1.DBD0, 1 s
   "84_Setpoints_E600_CB_HighHigh" : Real = PLC "84_Setpoints".E600_CB_HighHigh AT %DB1.DBD0, 1 s
   "84_Setpoints_FD001_Min" : Real = PLC "84_Setpoints".FD001_Min AT %DB1.DBD0, 1 s
   "84_Setpoints_PIT113_Pilot_Target(1)" : Real = PLC "62_Warning_Data".GCU_WARNING_WORD_01 AT %DB1.DBD0, 1 s
   "84_Setpoints_PIT205_Target(1)" : Real = PLC "84_Setpoints".PIT205_Target AT %DB1.DBD0, 1 s
   "84_Setpoints_E600_CB_Target" : Real = PLC "84_Setpoints".E600_CB_Target AT %DB1.DBD0, 1 s
   "84_Setpoints_E600_BWT_Target" : Real = PLC "84_Setpoints".E600_BWT_Target AT %DB1.DBD0, 1 s
   "86_Times_CV127_OPEN_TIME_#1" : Time = PLC "86_Times".CV127_OPEN_TIME_#1 AT %DB1.DBX0.0, 1 s
   "86_Times_CV127_CLOSED_TIME" : Time = PLC "86_Times".CV127_CLOSED_TIME AT %DB1.DBX0.0, 1 s
   "86_Times_CV127_OPEN_TIME_#2" : Time = PLC "86_Times".CV127_OPEN_TIME_#2 AT %DB1.DBX0.0, 1 s
   "86_Times_CV124_OPEN_TIME" : Time = PLC "86_Times".CV124_OPEN_TIME AT %DB1.DBX0.0, 1 s
   "86_Times_CV124_CLOSE_TIME_PRG" : Time = PLC "86_Times".CV124_CLOSE_TIME_PRG AT %DB1.DBX0.0, 1 s
   "86_Times_CV114_OPEN_TIME" : Time = PLC "86_Times".CV114_OPEN_TIME AT %DB1.DBX0.0, 1 s
   "86_Times_CV206_OPEN_TIME" : Time = PLC "86_Times".CV206_OPEN_TIME AT %DB1.DBX0.0, 1 s
   "86_Times_CV207_OPEN_TIME" : Time = PLC "86_Times".CV207_OPEN_TIME AT %DB1.DBX0.0, 1 s
   "86_Times_CV215_OPEN_TIME" : Time = PLC "86_Times".CV215_OPEN_TIME AT %DB1.DBX0.0, 1 s
   "86_Times_CV215_CLOSE_TIME_PRG" : Time = PLC "86_Times".CV215_CLOSE_TIME_PRG AT %DB1.DBX0.0, 1 s
   "86_Times_CV216_OPEN_TIME" : Time = PLC "86_Times".CV216_OPEN_TIME AT %DB1.DBX0.0, 1 s
   "86_Times_CV216_CLOSE_TIME_PRG" : Time = PLC "86_Times".CV216_CLOSE_TIME_PRG AT %DB1.DBX0.0, 1 s
   "86_Times_CV216_OPEN_TIME_PRG" : Time = PLC "86_Times".CV216_OPEN_TIME_PRG AT %DB1.DBX0.0, 1 s
   "86_Times_CV206_CLOSE_TIME" : Time = PLC "86_Times".CV206_CLOSE_TIME AT %DB1.DBX0.0, 1 s
   "86_Times_CV207_CLOSE_TIME" : Time = PLC "86_Times".CV207_CLOSE_TIME AT %DB1.DBX0.0, 1 s
   "86_Times_CV114_CLOSE_TIME" : Time = PLC "86_Times".CV114_CLOSE_TIME AT %DB1.DBD0, 1 s
   "86_Times_CV215_CLOSE_TIME" : Time = PLC "86_Times".CV215_CLOSE_TIME AT %DB1.DBD0, 1 s
   "86_Times_CV216_CLOSE_TIME" : Time = PLC "86_Times".CV216_CLOSE_TIME AT %DB1.DBD0, 1 s
   "86_Times_CV124_CLOSE_TIME" : Time = PLC "86_Times".CV124_CLOSE_TIME AT %DB1.DBD0, 1 s
   "86_Times_X001_MAX_RUN_TIME" : Time = PLC "86_Times".X001_MAX_RUN_TIME AT %DB1.DBD0, 1 s
   "86_Times_X001_RUN_CNF_TIME" : Time = PLC "86_Times".X001_RUN_CNF_TIME AT %DB1.DBD0, 1 s
   "86_Times_FD_DET_DELAY" : Time = PLC "86_Times".FD_DET_DELAY AT %DB1.DBD0, 1 s
   "86_Times_FD_VRFCTN_TIME" : Time = PLC "86_Times".FD_VRFCTN_TIME AT %DB1.DBD0, 1 s
   "86_Times_FDU_DET_TIME" : Time = PLC "86_Times".FDU_DET_TIME AT %DB1.DBD0, 1 s
   "86_Times_MAX_IGNTN_SEQ_TIME" : Time = PLC "86_Times".MAX_IGNTN_SEQ_TIME AT %DB1.DBD0, 1 s
   "86_Times_MAX_MAIN_BURN_SEQ_TIME" : Time = PLC "86_Times".MAX_MAIN_BURN_SEQ_TIME AT %DB1.DBD0, 1 s
   "86_Times_MAX_PILOT_PURGE_SEQ_TIME" : Time = PLC "86_Times".MAX_PILOT_PURGE_SEQ_TIME AT %DB1.DBD0, 1 s
   "86_Times_O2_CHECK_TIME" : Time = PLC "86_Times".O2_CHECK_TIME AT %DB1.DBD0, 1 s
   "86_Times_STEP_MAX_TIME_STP_001(1)" : Time = PLC "86_Times".STEP_MAX_TIME_STP_001 AT %DB1.DBW0, 1 s
   "86_Times_STEP_MAX_TIME_STP_005(1)" : Time = PLC "86_Times".STEP_MAX_TIME_STP_005 AT %DB1.DBW0, 1 s